TYPE MAC_TrimmingDeck_HMW :
STRUCT
   xEnableControlWidth : BOOL;   // Enable control cap width in automatic {x|x|x|x|O}
   xDisableControlWidth : BOOL;   // Disable control cap width in automatic {x|x|x|x|O}
   xEnableControlWander : BOOL;   // Enable control cap wander in automatic {x|x|x|x|O}
   xDisableControlWander : BOOL;   // Disable control cap wander in automatic {x|x|x|x|O}
   xResetOffset : BOOL;   // Reset all trimming deck offset {x|x|x|x|O}
   xPresetOpSide : BOOL;   // Preset request operator side {x|x|x|x|M}
   xPresetOppOpSide : BOOL;   // Preset request opposite operator side {x|x|x|x|M}
   xEnableDisableCulletEdge : BOOL;   // Enable/Disable cullet edges trimming {x|x|x|x|O}
   xEnableOpeningOnCleaning : BOOL;   // Enable opening trimming deck on cleaning mode {x|x|x|x|O}
   xDisableOpeningOnCleaning : BOOL;   // Disable pening trimming deck on cleaning mode {x|x|x|x|O}
   dOffsetOpSide_cmm : DINT;   // Trimming deck offset to add operator side [mm/100] {mm/100|mm|-150|150|O}
   dPositionManCmdOpSide_cmm : DINT;   // Trimming deck manual position operator side [mm/100] {mm/100|mm|-150|150|O}
   dOffsetOppOpSide_cmm : DINT;   // Trimming deck offset to add opposite operator side [mm/100] {mm/100|mm|-150|150|O}
   dPositionManCmdOppOpSide_cmm : DINT;   // Trimming deck manual position opposite operator side [mm/100] {mm/100|mm|-150|150|O}
   rgxMan : MAC_TrimmingDeck_HMWR_Man;   // Manual commands {x|x|x|x|O}
END_STRUCT
END_TYPE

TYPE MAC_TrimmingDeck_HMWR_Man :
STRUCT
   x0 : BOOL;   // Operator side - Move to External
   x1 : BOOL;   // Operator side - Move to Internal
   x2 : BOOL;
   x3 : BOOL;
   x4 : BOOL;   // Opposite operator side - Move to External
   x5 : BOOL;   // Opposite operator side - Move to Internal
   x6 : BOOL;
   x7 : BOOL;
   x8 : BOOL;   // Both sides - Move to operator side
   x9 : BOOL;   // Both sides - Move to opposite operator side
   x10 : BOOL;
   x11 : BOOL;
   x12 : BOOL;   // Operator side - Move to External (Maintenance)
   x13 : BOOL;   // Operator side - Move to Internal (Maintenance)
   x14 : BOOL;
   x15 : BOOL;
   x16 : BOOL;   // Opposite operator side - Move to External (Maintenance)
   x17 : BOOL;   // Opposite operator side - Move to Internal (Maintenance)
   x18 : BOOL;
   x19 : BOOL;
   x20 : BOOL;   // Operator side - Positioning Command
   x21 : BOOL;   // Opposite operator side - Positioning Command
   x22 : BOOL;
   x23 : BOOL;
   x24 : BOOL;
   x25 : BOOL;
   x26 : BOOL;
   x27 : BOOL;
   x28 : BOOL;
   x29 : BOOL;
   x30 : BOOL;
   x31 : BOOL;
END_STRUCT
END_TYPE

TYPE MAC_TrimmingDeck_IN_MOTION :
STRUCT
   DR_MAJ_M : MOTION_INSTRUCTION[2];   // Drive jog
   DR_MAM_M : MOTION_INSTRUCTION[2];   // Drive positioning
   DR_MAS_M : MOTION_INSTRUCTION[2];   // Drive stop
END_STRUCT
END_TYPE

TYPE MAC_TrimmingDeck_OUT_MOTION :
STRUCT
   DR_MSO_M : MOTION_INSTRUCTION[2];   // Drive ON
   DR_MSF_M : MOTION_INSTRUCTION[2];   // Drive OFF
   DR_MASR_M : MOTION_INSTRUCTION[2];   // Drive reset faults
   DR_MAJ_M : MOTION_INSTRUCTION[2];   // Drive jog
   DR_MAM_M : MOTION_INSTRUCTION[2];   // Drive positioning
   DR_MCD_M : MOTION_INSTRUCTION[2];   // Drive change speed
   DR_MAS_M : MOTION_INSTRUCTION[2];   // Drive stop
   DR_MAH_M : MOTION_INSTRUCTION[2];   // Drive homing
END_STRUCT
END_TYPE

TYPE MAC_TrimmingDeck_PH :
STRUCT
   x0 : BOOL;   // Trimming deck moving
   x1 : BOOL;
   x2 : BOOL;
   x3 : BOOL;
   x4 : BOOL;
   x5 : BOOL;
   x6 : BOOL;
   x7 : BOOL;   // Trimming deck wait arming completed
   x8 : BOOL;
   x9 : BOOL;
   x10 : BOOL;
   x11 : BOOL;
   x12 : BOOL;
   x13 : BOOL;
   x14 : BOOL;
   x15 : BOOL;
   x16 : BOOL;
   x17 : BOOL;
   x18 : BOOL;
   x19 : BOOL;
   x20 : BOOL;
   x21 : BOOL;
   x22 : BOOL;
   x23 : BOOL;
   x24 : BOOL;
   x25 : BOOL;
   x26 : BOOL;
   x27 : BOOL;
   x28 : BOOL;
   x29 : BOOL;
   x30 : BOOL;
   x31 : BOOL;
END_STRUCT
END_TYPE

TYPE MAC_TrimmingDeckUpdate :
STRUCT
   ST_xIndexCons : BOOL;   // Index consistent
   PH_xPlateHooked : BOOL;   // PH Plate hooked
   OS_xPlateInWindows : BOOL;   // OS Plate in windows
   OF_xPlateInWindows : BOOL;   // OF Plate in windows
   OSR_xPlateInWindows : BOOL;   // OSR Plate in windows
   OSF_xPlateInWindows : BOOL;   // OSF Plate in windows
   OSR_xPlateOutHooked : BOOL;   // OSR Plate hooked
   OS_xPlateOutHooked : BOOL;   // OS Plate hooked
   tSearchPlate : GP_TrackingSearchPlate_STC;   // Search plate data
   AUX_dIDMemory : DINT;   // ID Memory
   AUX_dReaction_cmm : DINT;   // Reation space [mm/100]
   AUX_dPositionDecision_cmm : DINT;   // Decision position [mm/100]
   AUX_dPositionStopSearch_cmm : DINT;   // Stop search position [mm/100]
   AUX_dPositionStopHooked_cmm : DINT;   // Stop hooked position [mm/100]
   AUX_dIndex : DINT;   // Index
END_STRUCT
END_TYPE

TYPE MAC_TrimmingWheels :
STRUCT
   CONF_dTrimWheelCodeOpt : DINT;   // Trimming wheels pair number for optimizer [Num]
   CONF_dPositionWheel_cmm : DINT;   // Distance from the beggining (From origin to split line) [mm/100]
   CONF_dConveyorLength_cmm : DINT;   // Conveyor length [mm/100]
   CONF_dConveyorStopPos_cmm : DINT;   // Conveyor stop position (If -1 then no stop available) [mm/100]
   CONF_dAvailableSpaceToStop_cmm : DINT;   // Space available for stop glass on trim wheel [mm/100]
   CONF_dMaxLengthWorkable_cmm : DINT;   // Maximum plate length to stop on conveyor [mm/100]
   CONF_dTolerance_cmm : DINT[2];   // Trimming wheel tolerance [mm/100]
   CONF_dTrimWheelArmPos_cmm : DINT[2];   // Trimming wheel position to start arming [mm/100]
   CONF_dStopCamPos_cmm : DINT[2];   // Trimming wheel position stop cam [mm/100]
   CONF_dSlowDownPos_cmm : DINT[2];   // Trimming wheels position slow down [mm/100]
   CONF_dTrimWheelHomePos_cmm : DINT[2];   // Trimming wheel home position [mm/100]
   CONF_dTrimWheelHomeSensorPos_cmm : DINT[2];   // Trimming wheel sensor home position [mm/100]
   CONF_dMaxTimeToReachPosition_ms : DINT[2];   // Maximum time to reach position [ms]
   CONF_dTrimWheelPreset : DINT[2];   // Trimming wheel preset encoder [pulse]
   CONF_dTrimWheelPresetZero_cmm : DINT[2];   // Trimming wheel encoder value in zero position [mm/100]
   CONF_dTrimWheelTargetWindow_cmm : DINT[2];   // Trimming wheel tollerance window on request position [mm/100]
   CONF_dTrimWheelDecWindow_cmm : DINT[2];   // Trimming wheel tollerance window on deceleration position [mm/100]
   CONF_dTrimWheelCleanPos_cmm : DINT[2];   // Trimming wheel cleaning position [mm/100]
   CONF_dTrimWheelMinPos_cmm : DINT[2];   // Trimming wheel minimum position [mm/100]
   CONF_dTrimWheelMaxPos_cmm : DINT[2];   // Trimming wheel maximum position [mm/100]
   CONF_dTrimWheelMinRange_cmm : DINT[2];   // Trimming wheel minimum work range [mm/100]
   CONF_dTrimWheelMaxRange_cmm : DINT[2];   // Trimming wheel maximum work range [mm/100]
   CONF_dSlowDownSpeed_mm_min : DINT[2];   // Trimming wheel slow down speed [mm/min]
   CONF_dSearchHomeSpeed_mm_min : DINT[2];   // Search home speed [mm/min]
   CONF_dAutoSpeed_mm_min : DINT[2];   // Trimming wheel automatic speed [mm/min]
   CONF_dManualSpeed_mm_min : DINT[2];   // Trimming wheel manual speed [mm/min]
   CONF_rTrimWheelPresetScaling : REAL[2];   // Trimming wheel preset scaling [(mm/100) / pulse]
   CONF_rAcceleration_m_s2 : REAL[2];   // Trimming wheel acceleration ramp [m/s2]
   CONF_rDeceleration_m_s2 : REAL[2];   // Trimming wheel deceleration ramp [m/s2]
   ST_xReqStartOpSide : BOOL;   // Request start operator side
   ST_xReqAbortOpSide : BOOL;   // Request abort operator side
   ST_xReqResetOffsetOpSide : BOOL;   // Request reset offset operator side
   ST_xReqStartTranslationOpSide : BOOL;   // Request start for translation operator side
   ST_xReqAbortTranslationOpSide : BOOL;   // Request abort for translation operator side
   ST_xReqResetOffsetTranslationOpSide : BOOL;   // Request reset offset for translation operator side
   ST_xReqUpdateTargetTranslationOpSide : BOOL;   // Request update target for translation operator side
   ST_xReqStartOppOpSide : BOOL;   // Request start opposite operator side
   ST_xReqAbortOppOpSide : BOOL;   // Request abort opposite operator side
   ST_xReqResetOffsetOppOpSide : BOOL;   // Request reset offset opposite operator side
   ST_xReqStartTranslationOppOpSide : BOOL;   // Request start for translation opposite operator side
   ST_xReqAbortTranslationOppOpSide : BOOL;   // Request abort for translation opposite operator side
   ST_xReqResetOffsetTranslationOppOpSide : BOOL;   // Request reset offset for translation opposite operator side
   ST_xReqUpdateTargetTranslationOppOpSide : BOOL;   // Request update target for translation opposite operator side
   ST_xReqResetOffsetGeneral : BOOL;   // Request reset offset general
   ST_xAxleHomedOpSide : BOOL;   // Axle homed operator side
   ST_xAxleHomedOppOpSide : BOOL;   // Axle homed opposite operator side
   ST_xTailBreakOppOpSide : BOOL;   // Tail break opposite operator side
   ST_xInitialConditionOpSideOK : BOOL;   // Initial condition OK operator side
   ST_xConditionOKPhaseadvancementOpSide : BOOL;   // Condition OK phase advancement operator side
   ST_xInitialConditionOppOpSideOK : BOOL;   // Initial condition OK opposite operator side
   ST_xConditionOKPhaseadvancementOppOpSide : BOOL;   // Condition OK phase advancement opposite operator side
   ST_xCleaningConditionOK : BOOL;   // Cleaning condition OK
   ST_xStopMachineFaultOpSide : BOOL;   // Stopped machine faults operator side
   ST_xStopNextCycleFaultOpSide : BOOL;   // Stopped next cycle faults operator side
   ST_xStopMachineFaultOppOpSide : BOOL;   // Stopped machine faults opposite operator side
   ST_xStopNextCycleFaultOppOpSide : BOOL;   // Stopped next cycle faults opposite operator side
   ST_xConditionOKStopCycle : BOOL;   // Condition OK for stop cycle
   ST_xConditionForStayDownInStaticMode : BOOL;   // Condition OK for stay down in static mode
   ST_xOutputEnableOpSide : BOOL;   // Output enable operator side
   ST_xOutputEnableHomeOpSide : BOOL;   // Output enable for home cycle operator side
   ST_xMachineFaultOpSide : BOOL;   // Machine with faults operator side
   ST_xWarningFaultOpSide : BOOL;   // Machine with warnings operator side
   ST_xOutputEnableOppOpSide : BOOL;   // Output enable opposite operator side
   ST_xOutputEnableHomeOppOpSide : BOOL;   // Output enable for home cycle opposite operator side
   ST_xMachineFaultOppOpSide : BOOL;   // Machine with faults opposite operator side
   ST_xWarningFaultOppOpSide : BOOL;   // Machine with warnings opposite operator side
   ST_xPhasesInProgressOpSide : BOOL;   // Operator side wheel phase in progress
   ST_xPhasesInProgressOppOpSide : BOOL;   // Opposite operator side wheel phase in progress
   ST_xHeadPresence : BOOL;   // Head presence on conveyor
   ST_xTailPresence : BOOL;   // Tail presence on conveyor
   ST_xEnableControlError : BOOL;   // Enable control error
   ST_xConvoyInProgress : BOOL;   // Convoy in progress
   ST_xFirstCapInConv : BOOL;   // First plate in convoy
   ST_xQualityInProgress : BOOL;   // Quality plate in progress
   ST_xCulletInProgress : BOOL;   // Cullet plate in progress
   ST_xInWorkOpSide : BOOL;   // Trimming wheel in work operator side
   ST_xInWorkOppOpSide : BOOL;   // Trimming wheel in work opposite operator side
   ST_xOutsideLimitFWOpSide : BOOL;   // Trimming wheel outside limit FW operator side
   ST_xOutsideLimitFWOppOpSide : BOOL;   // Trimming wheel outside limit FW opposite operator side
   ST_xOutsideLimitBWOpSide : BOOL;   // Trimming wheel outside limit BW operator side
   ST_xOutsideLimitBWOppOpSide : BOOL;   // Trimming wheel outside limit BW opposite operator side
   ST_xSafetyMovementOpSide : BOOL;   // Trimming wheel safety movement operator side
   ST_xSafetyMovementOppOpSide : BOOL;   // Trimming wheel safety movement opposite operator side
   ST_xFiringOpSide : BOOL;   // Firing trimming wheel operator side
   ST_xFiringOppOpSide : BOOL;   // Firing trimming wheel opposite operator side
   ST_xManualTrimEdgeOpSide : BOOL;   // Manual trimming edge operator side
   ST_xManualTrimEdgeOppOpSide : BOOL;   // Manual trimming edge opposite operator side
   ST_xInPositionOpSide : BOOL;   // Wheel in position operator side
   ST_xInPositionOppOpSide : BOOL;   // Wheel in position opposite operator side
   ST_xInSlowDownOpSide : BOOL;   // Wheel in slow down operator side
   ST_xInSlowDownOppOpSide : BOOL;   // Wheel in slow down opposite operator side
   ST_xInStopCamPositionOpSide : BOOL;   // Wheel in stop cam position operator side
   ST_xInStopCamPositionOppOpSide : BOOL;   // Wheel in stop cam position opposite operator side
   ST_xInStopCamManualOpSide : BOOL;   // Wheel in manual stop cam operator side
   ST_xInStopCamManualOppOpSide : BOOL;   // Wheel in manual stop cam opposite operator side
   ST_xInStopCamManualPositionOpSide : BOOL;   // Wheel in manual stop cam position operator side
   ST_xInStopCamManualPositionOppOpSide : BOOL;   // Wheel in manual stop cam position opposite operator side
   ST_xInSlowDownManualOpSide : BOOL;   // Wheel in manual slow down operator side
   ST_xInSlowDownManualOppOpSide : BOOL;   // Wheel in manual slow down opposite operator side
   ST_xInSlowDownManualPosOpSide : BOOL;   // Wheel in manual positioning slow down operator side
   ST_xInSlowDownManualPosOppOpSide : BOOL;   // Wheel in manual slow down positioning opposite operator side
   ST_xPositionReachedOpSide : BOOL;   // Wheel position reached operator side
   ST_xPositionReachedOppOpSide : BOOL;   // Wheel position reached opposite operator side
   ST_xInitialConditionHomeOpSide : BOOL;   // Initial condition for home cycle operator side
   ST_xInitialConditionHomeOppOpSide : BOOL;   // Initial condition for home cycle opposite operator side
   ST_xTailBreakOpSide : BOOL;   // Tail break operator side
   ST_xPreBreakingOpSide : BOOL;   // Wheel for pre breaking operator side
   ST_xPreBreakingOppOpSide : BOOL;   // Wheel for pre breaking opposite operator side
   ST_xPhaseONOpSide : BOOL;   // Wheel descent phase ON operator side
   ST_xPhaseONOppOpSide : BOOL;   // Wheel descent phase ON opposite operator side
   OSR_xStopConveyor : BOOL;   // OSR Stop conveyor
   OSR_xArmOpSide : BOOL;   // OSR Arming trimming wheel operator side
   OSR_xEndArmOpSide : BOOL;   // OSR End arming trimming wheel operator side
   OSR_xArmOppOpSide : BOOL;   // OSR Arming trimming wheel opposite operator side
   OSR_xEndArmOppOpSide : BOOL;   // OSR End arming trimming wheel opposite operator side
   OSR_xReqUpdateTargetTranslationOpSide : BOOL;   // OSR request update target for translation operator side
   OSR_xReqUpdateTargetTranslationOppOpSide : BOOL;   // OSR request update target for translation opposite operator side
   OSR_xStartPositioningOpSide : BOOL;   // OSR start positioning operator side
   OSR_xStartPositioningOppOpSide : BOOL;   // OSR start positioning opposite operator side
   OSR_xReqHomeCycleOpSide : BOOL;   // OSR Request home cycle operator side
   OSR_xReqHomeCycleOppOpSide : BOOL;   // OSR Request home cycle opposite operator side
   OSR_xIncrementOffsetOpSide : BOOL;   // OSR Increment offset operator side
   OSR_xDecrementOffsetOpSide : BOOL;   // OSR Decrement offset operator side
   OSR_xIncrementOffsetOppOpSide : BOOL;   // OSR Increment offset opposite operator side
   OSR_xDecrementOffsetOppOpSide : BOOL;   // OSR Decrement offset opposite operator side
   OS_xIncrementOffsetOpSide : BOOL;   // OS Increment offset operator side
   OS_xDecrementOffsetOpSide : BOOL;   // OS Decrement offset operator side
   OS_xIncrementOffsetOppOpSide : BOOL;   // OS Increment offset opposite operator side
   OS_xDecrementOffsetOppOpSide : BOOL;   // OS Decrement offset opposite operator side
   OSF_xFiringOpSide : BOOL;   // OSF Firing trimming wheel operator side
   OSF_xFiringOppOpSide : BOOL;   // OSF Firing trimming wheel opposite operator side
   OF_xFiringOpSide : BOOL;   // OF Firing trimming wheel operator side
   OF_xFiringOppOpSide : BOOL;   // OF Firing trimming wheel opposite operator side
   OS_xFiringOpSide : BOOL;   // OS Firing trimming wheel operator side
   OS_xFiringOppOpSide : BOOL;   // OS Firing trimming wheel opposite operator side
   OS_xStopConveyor : BOOL;   // OS Stop conveyor
   OS_xArmOpSide : BOOL;   // OS Arming trimming wheel operator side
   OS_xArmOppOpSide : BOOL;   // OS Arming trimming wheel opposite operator side
   OS_xReqUpdateTargetTranslationOpSide : BOOL;   // OS request update target for translation operator side
   OS_xReqUpdateTargetTranslationOppOpSide : BOOL;   // OS request update target for translation opposite operator side
   OS_xStartPositioningOpSide : BOOL;   // OS start positioning operator side
   OS_xStartPositioningOppOpSide : BOOL;   // OS start positioning opposite operator side
   OS_xReqHomeCycleOpSide : BOOL;   // OS Request home cycle operator side
   OS_xReqHomeCycleOppOpSide : BOOL;   // OS Request home cycle opposite operator side
   PH_xWaitPlateOpSide : BOOL;   // PH wait plate operator side
   PH_xWaitPlateOppOpSide : BOOL;   // PH wait plate opposite operator side
   PH_xFiringPlateOpSide : BOOL;   // PH firing operator side
   PH_xFiringPlateOppOpSide : BOOL;   // PH firing opposite operator side
   PH_xEndFiringPlateOpSide : BOOL;   // PH end firing operator side
   PH_xEndFiringPlateOppOpSide : BOOL;   // PH end firing opposite operator side
   PH_xPosTrOpSide : BOOL;   // PH translation positioning operator side
   PH_xPosTrOppOpSide : BOOL;   // PH translation positioning opposite operator side
   PH_xEndPosTrOpSide : BOOL;   // PH end translation positioning operator side
   PH_xEndPosTrOppOpSide : BOOL;   // PH end translation positioning opposite operator side
   PH_xReleaseSensorHomeOpSide : BOOL;   // PH Release sensor home operator side
   PH_xHomeCycleOpSide : BOOL;   // PH Home cycle operator side
   PH_xEndHomeCycleOpSide : BOOL;   // PH End Home cycle operator side
   PH_xReleaseSensorHomeOppOpSide : BOOL;   // PH Release sensor home opposite operator side
   PH_xHomeCycleOppOpSide : BOOL;   // PH Home cycle opposite operator side
   PH_xEndHomeCycleOppOpSide : BOOL;   // PH End Home cycle opposite operator side
   PH : MAC_TrimmingWheels_PH;   // Phases
   INPUT_xTrimDeckMoveInProgress : BOOL;   // Trimming deck moving in progress
   INPUT_xSBStopConveyor : BOOL;   // Stop conveyor on each plate
   INPUT_xSBSendToCullet : BOOL;   // Send to cullet
   INPUT_xSBSecondChoice : BOOL;   // Change destination to 2° Choice
   INPUT_xProtectionMotor : DINT;   // Motor protection
   INPUT_xLocalSafetySwitch : DINT;   // Local safety switch
   INPUT_xMotorThermalProbe : DINT;   // Motor Thermal Probe
   INPUT_xProtectionBrake : DINT;   // Brake protection
   INPUT_xBrakeFeedback : DINT;   // Brake feedback
   INPUT_xDriveInhibit : DINT;   // Drive inhibit
   INPUT_xDriveReady : DINT;   // Drive ready
   INPUT_xDriveError : DINT;   // Drive Error
   INPUT_xDriveFeedback : DINT;   // Drive Feedback
   INPUT_xDriveDeceleration : DINT;   // Drive deceleration
   INPUT_xHomePosition : DINT;   // Home position
   INPUT_xDriveHomedStatus : DINT;   // Drive homed status
   INPUT_xOverstrokeExternal : DINT;   // External overstroke
   INPUT_xOverstrokeInternal : DINT;   // Internal overstroke
   INPUT_xSBTrimWheelFastRise : DINT;   // Trimming wheel fast rise
   INPUT_xSBTrimWheelToCenterLine : DINT;   // Trimming wheel translation to center line
   INPUT_xSBTrimWheelToExternal : DINT;   // Trimming wheel translation to external
   INPUT_xSQTrimWheelHigh : DINT;   // Trimming wheel in high position
   INPUT_xSBTrimWheelDescent : DINT;   // Trimming wheel descending
   INPUT_xSBTrimWheelLift : DINT;   // Trimming wheel lifting
   INPUT_dRealSpeed_mm_min : DINT[2];   // Trimming wheel translation real speed [mm/min]
   INPUT_rAccDecRamp_m_s2 : REAL[2];   // Trimming wheel conveyor acceleration / decelaration ramp [m/s2]
   INPUT_dEncoder : DINT[2];   // Encoder pulse
   INPUT_dEncoderTranslation : DINT[2];   // Encoder pulse for translation
   OUTPUT_xSBStopConveyor : BOOL;   // Stop conveyor on each plate
   OUTPUT_xSBSendToCullet : BOOL;   // Send to cullet
   OUTPUT_xSBSecondChoice : BOOL;   // Change destination to 2° Choise
   OUTPUT_xDescent : DINT;   // Trimming wheel descending
   OUTPUT_xBlow : DINT;   // Trimming wheel blowing
   OUTPUT_xDriveReset : DINT;   // Drive reset faults
   OUTPUT_xDriveEnable : DINT;   // Output
   OUTPUT_xRun : DINT;   // Run
   OUTPUT_xReverse : DINT;   // Reverse
   OUTPUT_xPositioning : DINT;   // Positioning
   OUTPUT_xChangeSpeed : DINT;   // Change speed
   OUTPUT_xHoming : DINT;   // Homing
   OUTPUT_dEncoder : DINT[2];   // Encoder pulse
   OUTPUT_dEncoderTranslation : DINT[2];   // Encoder pulse for translation
   AUX_dOffsetGeneral_cmm : DINT;   // Offset translation for both wheel [mm/100]
   AUX_dReqLengthPlate_cmm : DINT[2];   // Request length plate [mm/100]
   AUX_dReqPositionPlate_cmm : DINT[2];   // Request plate position [mm/100]
   AUX_dReqTargetPosTranslation_cmm : DINT[2];   // Request target position translation [mm/100]
   AUX_dHeadPosition_cmm : DINT[2];   // Plate head position [mm/100]
   AUX_dTailPosition_cmm : DINT[2];   // Plate tail position [mm/100]
   AUX_dLengthPlate_cmm : DINT[2];   // Plate length [mm/100]
   AUX_dRampSpace_cmm : DINT[2];   // Ramp space [mm/100]
   AUX_dTrimWheelTarget_cmm : DINT[2];   // Trimming wheel target position without offset [mm/100]
   AUX_dCopyEncoderValue_cmm : DINT[2];   // Copy encoder value [mm/100]
   AUX_dPositionWheelBrk_cmm : DINT[2];   // Actual position of trimming wheel [mm/100]
   AUX_dDifferPositionBrkTailMode_cmm : DINT[2];   // Actual differ position tail break mode [mm/100]
   AUX_dActTransPosition_cmm : DINT[2];   // Actual translation position [mm/100]
   AUX_dOffsetSingle_cmm : DINT[2];   // Offset translation for single wheel [mm/100]
   AUX_dOffsetStep : DINT[2];   // Offset change for each step [mm/100]
   AUX_dFinalTarget_cmm : DINT[2];   // Final target [mm/100]
   AUX_dCopyValueEnc_cmm : DINT[2];   // Copy value encoder [mm/100]
   AUX_dCounterForAlarmEnc_cmm : DINT[2];   // Counter value for alarm encoder [mm/100]
   AUX_dReqSpeed_mm_min : DINT[2];   // Trimming deck requested speed [mm/min]
   AUX_dRealSpeed_mm_min : DINT[2];   // Trimming deck real speed [mm/min]
   AUX_dTotalCaps : DINT[2];   // Total caps coming for target
   AUX_rgxActivate : DINT[2];   // Activate action for convoy caps
   AUX_rgdConvoyGapsOpSide : DINT[3];   // Convoy gaps operator side [mm/100]
   AUX_rgdConvoyGapsOppOpSide : DINT[3];   // Convoy gaps operator side [mm/100]
   AUX_rgdConvoyLengthsOpSide : DINT[4];   // Convoy cap lengths operator side [mm/100]
   AUX_rgdConvoyLengthsOppOpSide : DINT[4];   // Convoy cap lengths operator side [mm/100]
   AUX_dSearchPlateDataOpSide : UDT_SearchPlateAuxData;   // Auxiliary data for searching plate operator side
   AUX_dSearchPlateDataOppOpSide : UDT_SearchPlateAuxData;   // Auxiliary data for searching plate opposite operator side
   AUX_dSearchPlateDataTranslationOpSide : UDT_SearchPlateAuxData;   // Auxiliary data for searching plate for translation operator side
   AUX_dSearchPlateDataTranslationOppOpSide : UDT_SearchPlateAuxData;   // Auxiliary data for searching plate for translation opposite operator side
   tmON_RequestHomeCycle : TIMER[2];   // Request home cycle
   tmON_EncPreset : TIMER[2];   // Encoder preset
   tmON_CheckEncoderTimeOut : TIMER[2];   // Check encoder time out
   tmON_TrimWheelTimeOut : TIMER[2];   // Trimming wheels time out
   tmON_TrimWheelBlow : TIMER[2];   // Trimming wheels blow time
   tmON_Wait : TIMER[2];   // Wait for glass process
   tmOF_DriveEnable : TIMER[2];   // Drive enable timer
   tmON_FeedbackTimeOut : TIMER[2];   // Feedback time out
   tmON_BrakeFeedbackTimeOut : TIMER[2];   // Brake feedback time out
   tmON_FeedbackDriveReady : TIMER[2];   // Drive ready feedback timer
   tmON_ReadyToMoveDelay : TIMER[2];   // Drive ready to move timer
   tmOF_DelayOnChangeDirection : TIMER[4];   // Delay on change direction
END_STRUCT
END_TYPE

TYPE MAC_TrimmingWheels_ALM :
STRUCT
   rgxStoppingFault : MAC_TrimmingWheels_ALM_SF[1];   // Generic stopping faults
   rgxFault : MAC_TrimmingWheels_ALM_F[1];   // Generic faults
   rgxWarning : MAC_TrimmingWheels_ALM_W[1];   // Generic warning
END_STRUCT
END_TYPE

TYPE MAC_TrimmingWheels_ALM_F :
STRUCT
   x0 : BOOL;   // Trimming wheel position error operator side
   x1 : BOOL;
   x2 : BOOL;
   x3 : BOOL;
   x4 : BOOL;
   x5 : BOOL;
   x6 : BOOL;
   x7 : BOOL;
   x8 : BOOL;
   x9 : BOOL;
   x10 : BOOL;   // Trimming wheel position error opposite operator side
   x11 : BOOL;
   x12 : BOOL;
   x13 : BOOL;
   x14 : BOOL;
   x15 : BOOL;
   x16 : BOOL;
   x17 : BOOL;
   x18 : BOOL;
   x19 : BOOL;
   x20 : BOOL;
   x21 : BOOL;
   x22 : BOOL;
   x23 : BOOL;
   x24 : BOOL;
   x25 : BOOL;
   x26 : BOOL;
   x27 : BOOL;
   x28 : BOOL;
   x29 : BOOL;
   x30 : BOOL;
   x31 : BOOL;
END_STRUCT
END_TYPE

TYPE MAC_TrimmingWheels_ALM_SF :
STRUCT
   x0 : BOOL;   // Trimming wheel protection motor operator side
   x1 : BOOL;   // Trimming wheel drive error operator side
   x2 : BOOL;   // Trimming wheel drive feedback error operator side
   x3 : BOOL;   // Trimming wheel protection brake operator side
   x4 : BOOL;   // Trimming wheel brake feedback error operator side
   x5 : BOOL;
   x6 : BOOL;
   x7 : BOOL;
   x8 : BOOL;
   x9 : BOOL;
   x10 : BOOL;   // Trimming wheel protection motor opposite operator side
   x11 : BOOL;   // Trimming wheel drive error opposite operator side
   x12 : BOOL;   // Trimming wheel drive feedback error opposite operator side
   x13 : BOOL;   // Trimming wheel protection brake opposite operator side
   x14 : BOOL;   // Trimming wheel brake feedback error opposite operator side
   x15 : BOOL;
   x16 : BOOL;
   x17 : BOOL;
   x18 : BOOL;
   x19 : BOOL;
   x20 : BOOL;
   x21 : BOOL;
   x22 : BOOL;
   x23 : BOOL;
   x24 : BOOL;
   x25 : BOOL;
   x26 : BOOL;
   x27 : BOOL;
   x28 : BOOL;
   x29 : BOOL;
   x30 : BOOL;
   x31 : BOOL;
END_STRUCT
END_TYPE

TYPE MAC_TrimmingWheels_ALM_W :
STRUCT
   x0 : BOOL;
   x1 : BOOL;
   x2 : BOOL;
   x3 : BOOL;
   x4 : BOOL;
   x5 : BOOL;
   x6 : BOOL;
   x7 : BOOL;
   x8 : BOOL;
   x9 : BOOL;
   x10 : BOOL;
   x11 : BOOL;
   x12 : BOOL;
   x13 : BOOL;
   x14 : BOOL;
   x15 : BOOL;
   x16 : BOOL;
   x17 : BOOL;
   x18 : BOOL;
   x19 : BOOL;
   x20 : BOOL;
   x21 : BOOL;
   x22 : BOOL;
   x23 : BOOL;
   x24 : BOOL;
   x25 : BOOL;
   x26 : BOOL;
   x27 : BOOL;
   x28 : BOOL;
   x29 : BOOL;
   x30 : BOOL;
   x31 : BOOL;
END_STRUCT
END_TYPE

TYPE MAC_TrimmingWheels_HMR :
STRUCT
   xStopConveyorEnabled : BOOL;   // Stop conveyor on each plate enabled {x|x|x|x|O}
   xAutoTrim : BOOL;   // Trimming wheel in auto mode {x|x|x|x|O}
   xDynamicTrim : BOOL;   // Trimming wheel in dynamic mode {x|x|x|x|O}
   xBlowChipsEnabled : BOOL;   // Trimming wheel blow chips enabled {x|x|x|x|O}
   xEnabledOpSide : BOOL;   // Trimming wheel operator side enabled {x|x|x|x|O}
   xEnabledOppOpSide : BOOL;   // Trimming wheel opposite operator side enabled {x|x|x|x|O}
   xManualCommandEnabled : BOOL;   // Trimming wheels manual command enabled {x|x|x|x|O}
   xWheelDownOpSide : BOOL;   // Trimming wheel down operator side {x|x|x|x|O}
   xWheelDownOppOpSide : BOOL;   // Trimming wheel down opposite operator side {x|x|x|x|O}
   rgdTarget_cmm : DINT[2];   // Trimming wheel request position [mm/100] {mm/100|mm|x|x|O}
   rgdPosition_cmm : DINT[2];   // Trimming wheel actual position [mm/100] {mm/100|mm|x|x|O}
   rgdState : DINT[2];   // Trimming wheel state (1=Rest position, 3=Run forward, 4=Run backward, 7=Alarm) {x|x|x|x|O}
   rgdEncoderPosition_cmm : DINT[2];   // Trimming wheel encoder position [mm/100] {mm/100|mm|x|x|O}
   rgdOffsetSingle_cmm : DINT[2];   // Trimming wheel offset single [mm/100] {mm/100|mm|-500|500|O}
   rgdOffsetDouble_cmm : DINT[2];   // Trimming wheel offset double [mm/100] {mm/100|mm|-500|500|O}
   rgdFinalTarget_cmm : DINT[2];   // Trimming wheel request position with offset [mm/100] {mm/100|mm|x|x|O}
   rgxMan : MAC_TrimmingWheels_HMWR_Man;   // Manual commands {x|x|x|x|O}
END_STRUCT
END_TYPE

TYPE MAC_TrimmingWheels_HMW :
STRUCT
   xEnableStopConveyor : BOOL;   // Enable stop conveyor {x|x|x|x|O}
   xDisableStopConveyor : BOOL;   // Disable stop conveyor {x|x|x|x|O}
   xReqAutoTrim : BOOL;   // Request automatic mode {x|x|x|x|O}
   xReqManualTrim : BOOL;   // Request manual mode {x|x|x|x|O}
   xReqDynamicTrim : BOOL;   // Request dynamic mode {x|x|x|x|O}
   xReqStaticTrim : BOOL;   // Request static mode {x|x|x|x|O}
   xReqOpSideTrimEdgeON : BOOL;   // Request descent for trimming edge operator side {x|x|x|x|O}
   xReqOpSideTrimEdgeOFF : BOOL;   // Request lifting for trimming edge operator side {x|x|x|x|O}
   xReqOppOpSideTrimEdgeON : BOOL;   // Request descent for trimming edge opposite operator side {x|x|x|x|O}
   xReqOppOpSideTrimEdgeOFF : BOOL;   // Request lifting for trimming edge opposite operator side {x|x|x|x|O}
   xEnableOpSide : BOOL;   // Enable trimming wheel operator side {x|x|x|x|O}
   xDisableOpSide : BOOL;   // Disable trimming wheel operator side {x|x|x|x|O}
   xEnableOppOpSide : BOOL;   // Enable trimming wheel opposite operator side {x|x|x|x|O}
   xDisableOppOpSide : BOOL;   // Disable trimming wheel opposite operator side {x|x|x|x|O}
   xEnableDisableBlowChips : BOOL;   // Enable/Disable chips blow {x|x|x|x|O}
   xEnableDisableManualCommand : BOOL;   // Enable/Disable manual command {x|x|x|x|O}
   xResetOffsetOpSide : BOOL;   // Reset all trimming wheel offset operator side {x|x|x|x|O}
   xResetOffsetOppOpSide : BOOL;   // Reset all trimming wheel offset opposite operator side {x|x|x|x|O}
   xPresetOpSide : BOOL;   // Preset request operator side {x|x|x|x|M}
   xPresetOppOpSide : BOOL;   // Preset request opposite operator side {x|x|x|x|M}
   xSemiAutoOpSide : BOOL;   // Operator side wheel in semi auto mode (Firing automatic and translation in manual) {x|x|x|x|O}
   xSemiAutoOppOpSide : BOOL;   // Opposite operator side wheel in semi auto mode (Firing automatic and translation in manual) {x|x|x|x|O}
   rgdBlowTime_ms : DINT[2];   // Blow time on trimming edge [ms] {ms|ms|0|5000|O}
   rgdOffsetStartTrim_cmm : DINT[2];   // Trimming wheels offset start trimming edge [mm/100] {mm/100|mm|-300|300|O}
   rgdOffsetStopTrim_cmm : DINT[2];   // Trimming wheels offset stop trimming edge [mm/100] {mm/100|mm|-300|300|O}
   rgdReactionTime_ms : DINT[2];   // Trimming wheel reaction time [ms] {ms|ms|0|5000|O}
   rgdOffsetPosition_cmm : DINT[2];   // Trimming wheel offset position [mm/100] {mm/100|mm|-150|150|O}
   rgdPlateLengthRise_perc : DINT[2];   // Trimming wheel percentage {x|x|0|100|O}
   rgdPositionManCmd_cmm : DINT[2];   // Trimming wheel manual position [mm/100] {mm/100|mm|0|500|O}
   rgxMan : MAC_TrimmingWheels_HMWR_Man;   // Manual commands {x|x|x|x|O}
END_STRUCT
END_TYPE

TYPE MAC_TrimmingWheels_HMWR_Man :
STRUCT
   x0 : BOOL;   // Trimming wheel descending operator side
   x1 : BOOL;   // Trimming wheel lifting operator side
   x2 : BOOL;   // Trimming wheel forward translation operator side
   x3 : BOOL;   // Trimming wheel backward translation operator side
   x4 : BOOL;   // Trimming wheel positioning operator side
   x5 : BOOL;   // Trimming wheel forward translation operator side (Maintenance Mode)
   x6 : BOOL;   // Trimming wheel backward translation operator side (Maintenance Mode)
   x7 : BOOL;
   x8 : BOOL;
   x9 : BOOL;
   x10 : BOOL;   // Trimming wheel descending opposite operator side
   x11 : BOOL;   // Trimming wheel lifting opposite operator side
   x12 : BOOL;   // Trimming wheel forward translation opposite operator side
   x13 : BOOL;   // Trimming wheel backward translation opposite operator side
   x14 : BOOL;   // Trimming wheel positioning opposite operator side
   x15 : BOOL;   // Trimming wheel forward translation opposite operator side (Maintenance Mode)
   x16 : BOOL;   // Trimming wheel backward translation opposite operator side (Maintenance Mode)
   x17 : BOOL;
   x18 : BOOL;
   x19 : BOOL;
   x20 : BOOL;
   x21 : BOOL;
   x22 : BOOL;
   x23 : BOOL;
   x24 : BOOL;
   x25 : BOOL;
   x26 : BOOL;
   x27 : BOOL;
   x28 : BOOL;
   x29 : BOOL;
   x30 : BOOL;
   x31 : BOOL;
END_STRUCT
END_TYPE
